   		OWF_Result[12].31:=0;
   	End_If;
   	If OWF_Input[5].[4] Then
   		OWF_Result[0]:=OWF_Result[0] + 1011754521+OWF_Add_c;
   		OWF_Add_c.0:=OWF_Result[0].31;
   		OWF_Result[0].31:=0;
   		OWF_Result[1]:=OWF_Result[1] + 1795510147+OWF_Add_c;
   		OWF_Add_c.1:=OWF_Result[1].31;
   		OWF_Result[1].31:=0;
   		OWF_Result[2]:=OWF_Result[2] + 543218634+OWF_Add_c;
   		OWF_Add_c.2:=OWF_Result[2].31;
   		OWF_Result[2].31:=0;
   		OWF_Result[3]:=OWF_Result[3] + 173475761+OWF_Add_c;
   		OWF_Add_c.3:=OWF_Result[3].31;
   		OWF_Result[3].31:=0;
   		OWF_Result[4]:=OWF_Result[4] + 535080772+OWF_Add_c;
   		OWF_Add_c.4:=OWF_Result[4].31;
   		OWF_Result[4].31:=0;
   		OWF_Result[5]:=OWF_Result[5] + 1289804735+OWF_Add_c;
   		OWF_Add_c.5:=OWF_Result[5].31;
   		OWF_Result[5].31:=0;
   		OWF_Result[6]:=OWF_Result[6] + 1812605489+OWF_Add_c;
   		OWF_Add_c.6:=OWF_Result[6].31;
   		OWF_Result[6].31:=0;
   		OWF_Result[7]:=OWF_Result[7] + 1203961891+OWF_Add_c;
   		OWF_Add_c.7:=OWF_Result[7].31;
   		OWF_Result[7].31:=0;
   		OWF_Result[8]:=OWF_Result[8] + 139150776+OWF_Add_c;
   		OWF_Add_c.8:=OWF_Result[8].31;
   		OWF_Result[8].31:=0;
   		OWF_Result[9]:=OWF_Result[9] + 1840895318+OWF_Add_c;
   		OWF_Add_c.9:=OWF_Result[9].31;
   		OWF_Result[9].31:=0;
   		OWF_Result[10]:=OWF_Result[10] + 576139644+OWF_Add_c;
   		OWF_Add_c.10:=OWF_Result[10].31;
   		OWF_Result[10].31:=0;
   		OWF_Result[11]:=OWF_Result[11] + 949700339+OWF_Add_c;
   		OWF_Add_c.11:=OWF_Result[11].31;
   		OWF_Result[11].31:=0;
   		OWF_Result[12]:=OWF_Result[12] + 707553602+OWF_Add_c;
   		OWF_Add_c.12:=OWF_Result[12].31;
   		OWF_Result[12].31:=0;
   	End_If;
   	If OWF_Input[5].[5] Then
   		OWF_Result[0]:=OWF_Result[0] + 341006670+OWF_Add_c;
   		OWF_Add_c.0:=OWF_Result[0].31;
   		OWF_Result[0].31:=0;
   		OWF_Result[1]:=OWF_Result[1] + 1545302097+OWF_Add_c;
   		OWF_Add_c.1:=OWF_Result[1].31;
   		OWF_Result[1].31:=0;
   		OWF_Result[2]:=OWF_Result[2] + 1059282447+OWF_Add_c;
   		OWF_Add_c.2:=OWF_Result[2].31;
   		OWF_Result[2].31:=0;
   		OWF_Result[3]:=OWF_Result[3] + 1918242377+OWF_Add_c;
   		OWF_Add_c.3:=OWF_Result[3].31;
   		OWF_Result[3].31:=0;
   		OWF_Result[4]:=OWF_Result[4] + 702854685+OWF_Add_c;
   		OWF_Add_c.4:=OWF_Result[4].31;
   		OWF_Result[4].31:=0;
   		OWF_Result[5]:=OWF_Result[5] + 1290612547+OWF_Add_c;
   		OWF_Add_c.5:=OWF_Result[5].31;
   		OWF_Result[5].31:=0;
   		OWF_Result[6]:=OWF_Result[6] + 1937985650+OWF_Add_c;
   		OWF_Add_c.6:=OWF_Result[6].31;
   		OWF_Result[6].31:=0;
   		OWF_Result[7]:=OWF_Result[7] + 1535904701+OWF_Add_c;
   		OWF_Add_c.7:=OWF_Result[7].31;
   		OWF_Result[7].31:=0;
   		OWF_Result[8]:=OWF_Result[8] + 57458357+OWF_Add_c;
   		OWF_Add_c.8:=OWF_Result[8].31;
   		OWF_Result[8].31:=0;
   		OWF_Result[9]:=OWF_Result[9] + 1270027244+OWF_Add_c;
   		OWF_Add_c.9:=OWF_Result[9].31;
   		OWF_Result[9].31:=0;
   		OWF_Result[10]:=OWF_Result[10] + 69146856+OWF_Add_c;
   		OWF_Add_c.10:=OWF_Result[10].31;
   		OWF_Result[10].31:=0;
   		OWF_Result[11]:=OWF_Result[11] + 1589075229+OWF_Add_c;
   		OWF_Add_c.11:=OWF_Result[11].31;
   		OWF_Result[11].31:=0;
   		OWF_Result[12]:=OWF_Result[12] + 458672961+OWF_Add_c;
   		OWF_Add_c.12:=OWF_Result[12].31;
   		OWF_Result[12].31:=0;
   	End_If;
   	If OWF_Input[5].[6] Then
   		OWF_Result[0]:=OWF_Result[0] + 1896310267+OWF_Add_c;
   		OWF_Add_c.0:=OWF_Result[0].31;
   		OWF_Result[0].31:=0;
   		OWF_Result[1]:=OWF_Result[1] + 1529180561+OWF_Add_c;
   		OWF_Add_c.1:=OWF_Result[1].31;
   		OWF_Result[1].31:=0;
   		OWF_Result[2]:=OWF_Result[2] + 2032481565+OWF_Add_c;
   		OWF_Add_c.2:=OWF_Result[2].31;
   		OWF_Result[2].31:=0;
   		OWF_Result[3]:=OWF_Result[3] + 537640111+OWF_Add_c;
   		OWF_Add_c.3:=OWF_Result[3].31;
   		OWF_Result[3].31:=0;
   		OWF_Result[4]:=OWF_Result[4] + 1272872794+OWF_Add_c;
   		OWF_Add_c.4:=OWF_Result[4].31;
   		OWF_Result[4].31:=0;
   		OWF_Result[5]:=OWF_Result[5] + 1539824454+OWF_Add_c;
   		OWF_Add_c.5:=OWF_Result[5].31;
   		OWF_Result[5].31:=0;
   		OWF_Result[6]:=OWF_Result[6] + 1430612137+OWF_Add_c;
   		OWF_Add_c.6:=OWF_Result[6].31;
   		OWF_Result[6].31:=0;
   		OWF_Result[7]:=OWF_Result[7] + 157560679+OWF_Add_c;
   		OWF_Add_c.7:=OWF_Result[7].31;
   		OWF_Result[7].31:=0;
   		OWF_Result[8]:=OWF_Result[8] + 259827156+OWF_Add_c;
   		OWF_Add_c.8:=OWF_Result[8].31;
   		OWF_Result[8].31:=0;
   		OWF_Result[9]:=OWF_Result[9] + 749936791+OWF_Add_c;
   		OWF_Add_c.9:=OWF_Result[9].31;
   		OWF_Result[9].31:=0;
   		OWF_Result[10]:=OWF_Result[10] + 1780248371+OWF_Add_c;
   		OWF_Add_c.10:=OWF_Result[10].31;
   		OWF_Result[10].31:=0;
   		OWF_Result[11]:=OWF_Result[11] + 1418315384+OWF_Add_c;
   		OWF_Add_c.11:=OWF_Result[11].31;
   		OWF_Result[11].31:=0;
   		OWF_Result[12]:=OWF_Result[12] + 406159660+OWF_Add_c;
   		OWF_Add_c.12:=OWF_Result[12].31;
   		OWF_Result[12].31:=0;
   	End_If;
   	If OWF_Input[5].[7] Then
   		OWF_Result[0]:=OWF_Result[0] + 2117716500+OWF_Add_c;
   		OWF_Add_c.0:=OWF_Result[0].31;
   		OWF_Result[0].31:=0;
   		OWF_Result[1]:=OWF_Result[1] + 1481111712+OWF_Add_c;
   		OWF_Add_c.1:=OWF_Result[1].31;
   		OWF_Result[1].31:=0;
   		OWF_Result[2]:=OWF_Result[2] + 1208238622+OWF_Add_c;
   		OWF_Add_c.2:=OWF_Result[2].31;
   		OWF_Result[2].31:=0;
   		OWF_Result[3]:=OWF_Result[3] + 1587378712+OWF_Add_c;
   		OWF_Add_c.3:=OWF_Result[3].31;
   		OWF_Result[3].31:=0;
   		OWF_Result[4]:=OWF_Result[4] + 1486187831+OWF_Add_c;
   		OWF_Add_c.4:=OWF_Result[4].31;
   		OWF_Result[4].31:=0;
   		OWF_Result[5]:=OWF_Result[5] + 1463632282+OWF_Add_c;
   		OWF_Add_c.5:=OWF_Result[5].31;
   		OWF_Result[5].31:=0;
   		OWF_Result[6]:=OWF_Result[6] + 594379430+OWF_Add_c;
   		OWF_Add_c.6:=OWF_Result[6].31;
   		OWF_Result[6].31:=0;
   		OWF_Result[7]:=OWF_Result[7] + 61907271+OWF_Add_c;
   		OWF_Add_c.7:=OWF_Result[7].31;
   		OWF_Result[7].31:=0;
   		OWF_Result[8]:=OWF_Result[8] + 1446292796+OWF_Add_c;
   		OWF_Add_c.8:=OWF_Result[8].31;
   		OWF_Result[8].31:=0;
   		OWF_Result[9]:=OWF_Result[9] + 1953507778+OWF_Add_c;
   		OWF_Add_c.9:=OWF_Result[9].31;
   		OWF_Result[9].31:=0;
   		OWF_Result[10]:=OWF_Result[10] + 1721398400+OWF_Add_c;
   		OWF_Add_c.10:=OWF_Result[10].31;
   		OWF_Result[10].31:=0;
   		OWF_Result[11]:=OWF_Result[11] + 704130819+OWF_Add_c;
   		OWF_Add_c.11:=OWF_Result[11].31;
   		OWF_Result[11].31:=0;
   		OWF_Result[12]:=OWF_Result[12] + 156099517+OWF_Add_c;
   		OWF_Add_c.12:=OWF_Result[12].31;
   		OWF_Result[12].31:=0;
   	End_If;
   	If OWF_Input[5].[8] Then
   		OWF_Result[0]:=OWF_Result[0] + 1443938657+OWF_Add_c;
   		OWF_Add_c.0:=OWF_Result[0].31;
   		OWF_Result[0].31:=0;
   		OWF_Result[1]:=OWF_Result[1] + 387077029+OWF_Add_c;
   		OWF_Add_c.1:=OWF_Result[1].31;
   		OWF_Result[1].31:=0;
   		OWF_Result[2]:=OWF_Result[2] + 331220417+OWF_Add_c;
   		OWF_Add_c.2:=OWF_Result[2].31;
   		OWF_Result[2].31:=0;
   		OWF_Result[3]:=OWF_Result[3] + 1153901105+OWF_Add_c;
   		OWF_Add_c.3:=OWF_Result[3].31;
   		OWF_Result[3].31:=0;
   		OWF_Result[4]:=OWF_Result[4] + 758718018+OWF_Add_c;
   		OWF_Add_c.4:=OWF_Result[4].31;
   		OWF_Result[4].31:=0;
   		OWF_Result[5]:=OWF_Result[5] + 1180469231+OWF_Add_c;
   		OWF_Add_c.5:=OWF_Result[5].31;
   		OWF_Result[5].31:=0;
   		OWF_Result[6]:=OWF_Result[6] + 451076221+OWF_Add_c;
   		OWF_Add_c.6:=OWF_Result[6].31;
   		OWF_Result[6].31:=0;
   		OWF_Result[7]:=OWF_Result[7] + 1957369555+OWF_Add_c;
   		OWF_Add_c.7:=OWF_Result[7].31;
   		OWF_Result[7].31:=0;
   		OWF_Result[8]:=OWF_Result[8] + 157679071+OWF_Add_c;
   		OWF_Add_c.8:=OWF_Result[8].31;
   		OWF_Result[8].31:=0;
   		OWF_Result[9]:=OWF_Result[9] + 999919265+OWF_Add_c;
   		OWF_Add_c.9:=OWF_Result[9].31;
   		OWF_Result[9].31:=0;
   		OWF_Result[10]:=OWF_Result[10] + 325782623+OWF_Add_c;
   		OWF_Add_c.10:=OWF_Result[10].31;
   		OWF_Result[10].31:=0;
   		OWF_Result[11]:=OWF_Result[11] + 1839549707+OWF_Add_c;
   		OWF_Add_c.11:=OWF_Result[11].31;
   		OWF_Result[11].31:=0;
   		OWF_Result[12]:=OWF_Result[12] + 210567637+OWF_Add_c;
   		OWF_Add_c.12:=OWF_Result[12].31;
   		OWF_Result[12].31:=0;
   	End_If;
   	If OWF_Input[5].[9] Then
   		OWF_Result[0]:=OWF_Result[0] + 1164800234+OWF_Add_c;
   		OWF_Add_c.0:=OWF_Result[0].31;
   		OWF_Result[0].31:=0;
   		OWF_Result[1]:=OWF_Result[1] + 373070247+OWF_Add_c;
   		OWF_Add_c.1:=OWF_Result[1].31;
   		OWF_Result[1].31:=0;
   		OWF_Result[2]:=OWF_Result[2] + 102655075+OWF_Add_c;
   		OWF_Add_c.2:=OWF_Result[2].31;
   		OWF_Result[2].31:=0;
   		OWF_Result[3]:=OWF_Result[3] + 1112504203+OWF_Add_c;
   		OWF_Add_c.3:=OWF_Result[3].31;
   		OWF_Result[3].31:=0;
   		OWF_Result[4]:=OWF_Result[4] + 728629506+OWF_Add_c;
   		OWF_Add_c.4:=OWF_Result[4].31;
   		OWF_Result[4].31:=0;
   		OWF_Result[5]:=OWF_Result[5] + 112310491+OWF_Add_c;
   		OWF_Add_c.5:=OWF_Result[5].31;
   		OWF_Result[5].31:=0;
   		OWF_Result[6]:=OWF_Result[6] + 1422404199+OWF_Add_c;
   		OWF_Add_c.6:=OWF_Result[6].31;
   		OWF_Result[6].31:=0;
   		OWF_Result[7]:=OWF_Result[7] + 1701166039+OWF_Add_c;
   		OWF_Add_c.7:=OWF_Result[7].31;
   		OWF_Result[7].31:=0;
   		OWF_Result[8]:=OWF_Result[8] + 2102782443+OWF_Add_c;
   		OWF_Add_c.8:=OWF_Result[8].31;
   		OWF_Result[8].31:=0;
   		OWF_Result[9]:=OWF_Result[9] + 1540134296+OWF_Add_c;
   		OWF_Add_c.9:=OWF_Result[9].31;
   		OWF_Result[9].31:=0;
   		OWF_Result[10]:=OWF_Result[10] + 2068205909+OWF_Add_c;
   		OWF_Add_c.10:=OWF_Result[10].31;
   		OWF_Result[10].31:=0;
   		OWF_Result[11]:=OWF_Result[11] + 1462437349+OWF_Add_c;
   		OWF_Add_c.11:=OWF_Result[11].31;
   		OWF_Result[11].31:=0;
   		OWF_Result[12]:=OWF_Result[12] + 1542204103+OWF_Add_c;
   		OWF_Add_c.12:=OWF_Result[12].31;
   		OWF_Result[12].31:=0;
   	End_If;
   	If OWF_Input[5].[10] Then
   		OWF_Result[0]:=OWF_Result[0] + 1094309781+OWF_Add_c;
   		OWF_Add_c.0:=OWF_Result[0].31;
   		OWF_Result[0].31:=0;
   		OWF_Result[1]:=OWF_Result[1] + 1799253283+OWF_Add_c;
   		OWF_Add_c.1:=OWF_Result[1].31;
   		OWF_Result[1].31:=0;
   		OWF_Result[2]:=OWF_Result[2] + 907784774+OWF_Add_c;
   		OWF_Add_c.2:=OWF_Result[2].31;
   		OWF_Result[2].31:=0;
   		OWF_Result[3]:=OWF_Result[3] + 1760595174+OWF_Add_c;
   		OWF_Add_c.3:=OWF_Result[3].31;
   		OWF_Result[3].31:=0;
   		OWF_Result[4]:=OWF_Result[4] + 1516380446+OWF_Add_c;
   		OWF_Add_c.4:=OWF_Result[4].31;
   		OWF_Result[4].31:=0;
   		OWF_Result[5]:=OWF_Result[5] + 525293244+OWF_Add_c;
   		OWF_Add_c.5:=OWF_Result[5].31;
   		OWF_Result[5].31:=0;
   		OWF_Result[6]:=OWF_Result[6] + 1469823607+OWF_Add_c;
   		OWF_Add_c.6:=OWF_Result[6].31;
   		OWF_Result[6].31:=0;
   		OWF_Result[7]:=OWF_Result[7] + 990094771+OWF_Add_c;
   		OWF_Add_c.7:=OWF_Result[7].31;
   		OWF_Result[7].31:=0;
   		OWF_Result[8]:=OWF_Result[8] + 206451193+OWF_Add_c;
   		OWF_Add_c.8:=OWF_Result[8].31;
   		OWF_Result[8].31:=0;
   		OWF_Result[9]:=OWF_Result[9] + 2094599626+OWF_Add_c;
   		OWF_Add_c.9:=OWF_Result[9].31;
   		OWF_Result[9].31:=0;
   		OWF_Result[10]:=OWF_Result[10] + 1804619518+OWF_Add_c;
   		OWF_Add_c.10:=OWF_Result[10].31;
   		OWF_Result[10].31:=0;
   		OWF_Result[11]:=OWF_Result[11] + 531327458+OWF_Add_c;
   		OWF_Add_c.11:=OWF_Result[11].31;
   		OWF_Result[11].31:=0;
   		OWF_Result[12]:=OWF_Result[12] + 914900243+OWF_Add_c;
   		OWF_Add_c.12:=OWF_Result[12].31;
   		OWF_Result[12].31:=0;
   	End_If;
   	If OWF_Input[5].[11] Then
   		OWF_Result[0]:=OWF_Result[0] + 1387671324+OWF_Add_c;
   		OWF_Add_c.0:=OWF_Result[0].31;
   		OWF_Result[0].31:=0;
   		OWF_Result[1]:=OWF_Result[1] + 770124107+OWF_Add_c;
   		OWF_Add_c.1:=OWF_Result[1].31;
   		OWF_Result[1].31:=0;
   		OWF_Result[2]:=OWF_Result[2] + 2104522684+OWF_Add_c;
   		OWF_Add_c.2:=OWF_Result[2].31;
   		OWF_Result[2].31:=0;
   		OWF_Result[3]:=OWF_Result[3] + 702616803+OWF_Add_c;
   		OWF_Add_c.3:=OWF_Result[3].31;
   		OWF_Result[3].31:=0;
   		OWF_Result[4]:=OWF_Result[4] + 453094356+OWF_Add_c;
   		OWF_Add_c.4:=OWF_Result[4].31;
   		OWF_Result[4].31:=0;
   		OWF_Result[5]:=OWF_Result[5] + 2109390133+OWF_Add_c;
   		OWF_Add_c.5:=OWF_Result[5].31;
   		OWF_Result[5].31:=0;
   		OWF_Result[6]:=OWF_Result[6] + 156781386+OWF_Add_c;
   		OWF_Add_c.6:=OWF_Result[6].31;
   		OWF_Result[6].31:=0;
   		OWF_Result[7]:=OWF_Result[7] + 1882451383+OWF_Add_c;
   		OWF_Add_c.7:=OWF_Result[7].31;
   		OWF_Result[7].31:=0;
   		OWF_Result[8]:=OWF_Result[8] + 1276007251+OWF_Add_c;
   		OWF_Add_c.8:=OWF_Result[8].31;
   		OWF_Result[8].31:=0;
   		OWF_Result[9]:=OWF_Result[9] + 1340635153+OWF_Add_c;
   		OWF_Add_c.9:=OWF_Result[9].31;
   		OWF_Result[9].31:=0;
   		OWF_Result[10]:=OWF_Result[10] + 225675392+OWF_Add_c;
   		OWF_Add_c.10:=OWF_Result[10].31;
   		OWF_Result[10].31:=0;
   		OWF_Result[11]:=OWF_Result[11] + 403241353+OWF_Add_c;
   		OWF_Add_c.11:=OWF_Result[11].31;
   		OWF_Result[11].31:=0;
   		OWF_Result[12]:=OWF_Result[12] + 1949018013+OWF_Add_c;
   		OWF_Add_c.12:=OWF_Result[12].31;
   		OWF_Result[12].31:=0;
   	End_If;
   	If OWF_Input[5].[12] Then
   		OWF_Result[0]:=OWF_Result[0] + 1384871639+OWF_Add_c;
   		OWF_Add_c.0:=OWF_Result[0].31;
   		OWF_Result[0].31:=0;
   		OWF_Result[1]:=OWF_Result[1] + 1594702713+OWF_Add_c;
   		OWF_Add_c.1:=OWF_Result[1].31;
   		OWF_Result[1].31:=0;
   		OWF_Result[2]:=OWF_Result[2] + 756803648+OWF_Add_c;
   		OWF_Add_c.2:=OWF_Result[2].31;
   		OWF_Result[2].31:=0;
   		OWF_Result[3]:=OWF_Result[3] + 26768879+OWF_Add_c;
   		OWF_Add_c.3:=OWF_Result[3].31;
   		OWF_Result[3].31:=0;
   		OWF_Result[4]:=OWF_Result[4] + 1679784822+OWF_Add_c;
   		OWF_Add_c.4:=OWF_Result[4].31;
   		OWF_Result[4].31:=0;
   		OWF_Result[5]:=OWF_Result[5] + 970059452+OWF_Add_c;
   		OWF_Add_c.5:=OWF_Result[5].31;
   		OWF_Result[5].31:=0;
   		OWF_Result[6]:=OWF_Result[6] + 1810393488+OWF_Add_c;
   		OWF_Add_c.6:=OWF_Result[6].31;
   		OWF_Result[6].31:=0;
   		OWF_Result[7]:=OWF_Result[7] + 488169811+OWF_Add_c;
   		OWF_Add_c.7:=OWF_Result[7].31;
   		OWF_Result[7].31:=0;
   		OWF_Result[8]:=OWF_Result[8] + 1304722861+OWF_Add_c;
   		OWF_Add_c.8:=OWF_Result[8].31;
   		OWF_Result[8].31:=0;
   		OWF_Result[9]:=OWF_Result[9] + 1892980786+OWF_Add_c;
   		OWF_Add_c.9:=OWF_Result[9].31;
   		OWF_Result[9].31:=0;
   		OWF_Result[10]:=OWF_Result[10] + 1092125948+OWF_Add_c;
   		OWF_Add_c.10:=OWF_Result[10].31;
   		OWF_Result[10].31:=0;
   		OWF_Result[11]:=OWF_Result[11] + 1982722541+OWF_Add_c;
   		OWF_Add_c.11:=OWF_Result[11].31;
   		OWF_Result[11].31:=0;
   		OWF_Result[12]:=OWF_Result[12] + 326633928+OWF_Add_c;
   		OWF_Add_c.12:=OWF_Result[12].31;
   		OWF_Result[12].31:=0;
   	End_If;
   	If OWF_Input[5].[13] Then
   		OWF_Result[0]:=OWF_Result[0] + 1000988417+OWF_Add_c;
   		OWF_Add_c.0:=OWF_Result[0].31;
   		OWF_Result[0].31:=0;
   		OWF_Result[1]:=OWF_Result[1] + 994193103+OWF_Add_c;
   		OWF_Add_c.1:=OWF_Result[1].31;
   		OWF_Result[1].31:=0;
   		OWF_Result[2]:=OWF_Result[2] + 1537710547+OWF_Add_c;
   		OWF_Add_c.2:=OWF_Result[2].31;
   		OWF_Result[2].31:=0;
   		OWF_Result[3]:=OWF_Result[3] + 15619081+OWF_Add_c;
   		OWF_Add_c.3:=OWF_Result[3].31;
   		OWF_Result[3].31:=0;
   		OWF_Result[4]:=OWF_Result[4] + 2143143663+OWF_Add_c;
   		OWF_Add_c.4:=OWF_Result[4].31;
   		OWF_Result[4].31:=0;
   		OWF_Result[5]:=OWF_Result[5] + 393950588+OWF_Add_c;
   		OWF_Add_c.5:=OWF_Result[5].31;
   		OWF_Result[5].31:=0;
   		OWF_Result[6]:=OWF_Result[6] + 1961783643+OWF_Add_c;
   		OWF_Add_c.6:=OWF_Result[6].31;
   		OWF_Result[6].31:=0;
   		OWF_Result[7]:=OWF_Result[7] + 2056947807+OWF_Add_c;
   		OWF_Add_c.7:=OWF_Result[7].31;
   		OWF_Result[7].31:=0;
   		OWF_Result[8]:=OWF_Result[8] + 939957448+OWF_Add_c;
   		OWF_Add_c.8:=OWF_Result[8].31;
   		OWF_Result[8].31:=0;
   		OWF_Result[9]:=OWF_Result[9] + 1853399300+OWF_Add_c;
   		OWF_Add_c.9:=OWF_Result[9].31;
   		OWF_Result[9].31:=0;
   		OWF_Result[10]:=OWF_Result[10] + 1339264557+OWF_Add_c;
   		OWF_Add_c.10:=OWF_Result[10].31;
   		OWF_Result[10].31:=0;
   		OWF_Result[11]:=OWF_Result[11] + 200481107+OWF_Add_c;
   		OWF_Add_c.11:=OWF_Result[11].31;
   		OWF_Result[11].31:=0;
   		OWF_Result[12]:=OWF_Result[12] + 1047995528+OWF_Add_c;
   		OWF_Add_c.12:=OWF_Result[12].31;
   		OWF_Result[12].31:=0;
   	End_If;
   	If OWF_Input[5].[14] Then
   		OWF_Result[0]:=OWF_Result[0] + 1208463242+OWF_Add_c;
   		OWF_Add_c.0:=OWF_Result[0].31;
   		OWF_Result[0].31:=0;
   		OWF_Result[1]:=OWF_Result[1] + 1623027587+OWF_Add_c;
   		OWF_Add_c.1:=OWF_Result[1].31;
   		OWF_Result[1].31:=0;
   		OWF_Result[2]:=OWF_Result[2] + 605083722+OWF_Add_c;
   		OWF_Add_c.2:=OWF_Result[2].31;
   		OWF_Result[2].31:=0;
   		OWF_Result[3]:=OWF_Result[3] + 1196976689+OWF_Add_c;
   		OWF_Add_c.3:=OWF_Result[3].31;
   		OWF_Result[3].31:=0;
   		OWF_Result[4]:=OWF_Result[4] + 2034493170+OWF_Add_c;
   		OWF_Add_c.4:=OWF_Result[4].31;
   		OWF_Result[4].31:=0;
   		OWF_Result[5]:=OWF_Result[5] + 718055369+OWF_Add_c;
   		OWF_Add_c.5:=OWF_Result[5].31;
   		OWF_Result[5].31:=0;
   		OWF_Result[6]:=OWF_Result[6] + 910332765+OWF_Add_c;
   		OWF_Add_c.6:=OWF_Result[6].31;
   		OWF_Result[6].31:=0;
   		OWF_Result[7]:=OWF_Result[7] + 1449925077+OWF_Add_c;
   		OWF_Add_c.7:=OWF_Result[7].31;
   		OWF_Result[7].31:=0;
   		OWF_Result[8]:=OWF_Result[8] + 839039994+OWF_Add_c;
   		OWF_Add_c.8:=OWF_Result[8].31;
   		OWF_Result[8].31:=0;
   		OWF_Result[9]:=OWF_Result[9] + 1168597276+OWF_Add_c;
   		OWF_Add_c.9:=OWF_Result[9].31;
   		OWF_Result[9].31:=0;
   		OWF_Result[10]:=OWF_Result[10] + 42917457+OWF_Add_c;
   		OWF_Add_c.10:=OWF_Result[10].31;
   		OWF_Result[10].31:=0;
   		OWF_Result[11]:=OWF_Result[11] + 1907752552+OWF_Add_c;
   		OWF_Add_c.11:=OWF_Result[11].31;
   		OWF_Result[11].31:=0;
   		OWF_Result[12]:=OWF_Result[12] + 1741695515+OWF_Add_c;
   		OWF_Add_c.12:=OWF_Result[12].31;
   		OWF_Result[12].31:=0;
   	End_If;
   	If OWF_Input[5].[15] Then
   		OWF_Result[0]:=OWF_Result[0] + 963845262+OWF_Add_c;
   		OWF_Add_c.0:=OWF_Result[0].31;
   		OWF_Result[0].31:=0;
   		OWF_Result[1]:=OWF_Result[1] + 1178480242+OWF_Add_c;
   		OWF_Add_c.1:=OWF_Result[1].31;
   		OWF_Result[1].31:=0;
   		OWF_Result[2]:=OWF_Result[2] + 555963648+OWF_Add_c;
   		OWF_Add_c.2:=OWF_Result[2].31;
   		OWF_Result[2].31:=0;
   		OWF_Result[3]:=OWF_Result[3] + 2035289100+OWF_Add_c;
   		OWF_Add_c.3:=OWF_Result[3].31;
   		OWF_Result[3].31:=0;
   		OWF_Result[4]:=OWF_Result[4] + 1602592723+OWF_Add_c;
   		OWF_Add_c.4:=OWF_Result[4].31;
   		OWF_Result[4].31:=0;
   		OWF_Result[5]:=OWF_Result[5] + 1321176695+OWF_Add_c;
   		OWF_Add_c.5:=OWF_Result[5].31;
   		OWF_Result[5].31:=0;
   		OWF_Result[6]:=OWF_Result[6] + 1370169932+OWF_Add_c;
   		OWF_Add_c.6:=OWF_Result[6].31;
   		OWF_Result[6].31:=0;
   		OWF_Result[7]:=OWF_Result[7] + 1543393295+OWF_Add_c;
   		OWF_Add_c.7:=OWF_Result[7].31;
   		OWF_Result[7].31:=0;
   		OWF_Result[8]:=OWF_Result[8] + 83738279+OWF_Add_c;
   		OWF_Add_c.8:=OWF_Result[8].31;
   		OWF_Result[8].31:=0;
   		OWF_Result[9]:=OWF_Result[9] + 725427957+OWF_Add_c;
   		OWF_Add_c.9:=OWF_Result[9].31;
   		OWF_Result[9].31:=0;
   		OWF_Result[10]:=OWF_Result[10] + 581206308+OWF_Add_c;
   		OWF_Add_c.10:=OWF_Result[10].31;
   		OWF_Result[10].31:=0;
   		OWF_Result[11]:=OWF_Result[11] + 491262647+OWF_Add_c;
   		OWF_Add_c.11:=OWF_Result[11].31;
   		OWF_Result[11].31:=0;
   		OWF_Result[12]:=OWF_Result[12] + 2147137437+OWF_Add_c;
   		OWF_Add_c.12:=OWF_Result[12].31;
   		OWF_Result[12].31:=0;
   	End_If;
   	If OWF_Input[5].[16] Then
   		OWF_Result[0]:=OWF_Result[0] + 2074453075+OWF_Add_c;
   		OWF_Add_c.0:=OWF_Result[0].31;
   		OWF_Result[0].31:=0;
   		OWF_Result[1]:=OWF_Result[1] + 108344464+OWF_Add_c;
   		OWF_Add_c.1:=OWF_Result[1].31;
   		OWF_Result[1].31:=0;
   		OWF_Result[2]:=OWF_Result[2] + 452532141+OWF_Add_c;
   		OWF_Add_c.2:=OWF_Result[2].31;
   		OWF_Result[2].31:=0;
   		OWF_Result[3]:=OWF_Result[3] + 1547961836+OWF_Add_c;
   		OWF_Add_c.3:=OWF_Result[3].31;
   		OWF_Result[3].31:=0;
   		OWF_Result[4]:=OWF_Result[4] + 1372224157+OWF_Add_c;
   		OWF_Add_c.4:=OWF_Result[4].31;
   		OWF_Result[4].31:=0;
   		OWF_Result[5]:=OWF_Result[5] + 1842815326+OWF_Add_c;
   		OWF_Add_c.5:=OWF_Result[5].31;
   		OWF_Result[5].31:=0;
   		OWF_Result[6]:=OWF_Result[6] + 614084210+OWF_Add_c;
   		OWF_Add_c.6:=OWF_Result[6].31;
   		OWF_Result[6].31:=0;
   		OWF_Result[7]:=OWF_Result[7] + 2105622125+OWF_Add_c;
   		OWF_Add_c.7:=OWF_Result[7].31;
   		OWF_Result[7].31:=0;
   		OWF_Result[8]:=OWF_Result[8] + 1347171274+OWF_Add_c;
   		OWF_Add_c.8:=OWF_Result[8].31;
   		OWF_Result[8].31:=0;
   		OWF_Result[9]:=OWF_Result[9] + 1124490238+OWF_Add_c;
   		OWF_Add_c.9:=OWF_Result[9].31;
   		OWF_Result[9].31:=0;
   		OWF_Result[10]:=OWF_Result[10] + 2064336718+OWF_Add_c;
   		OWF_Add_c.10:=OWF_Result[10].31;
   		OWF_Result[10].31:=0;
   		OWF_Result[11]:=OWF_Result[11] + 1049919562+OWF_Add_c;
   		OWF_Add_c.11:=OWF_Result[11].31;
   		OWF_Result[11].31:=0;
   		OWF_Result[12]:=OWF_Result[12] + 13830202+OWF_Add_c;
   		OWF_Add_c.12:=OWF_Result[12].31;
   		OWF_Result[12].31:=0;
   	End_If;
   	If OWF_Input[5].[17] Then
   		OWF_Result[0]:=OWF_Result[0] + 409887176+OWF_Add_c;
   		OWF_Add_c.0:=OWF_Result[0].31;
   		OWF_Result[0].31:=0;
   		OWF_Result[1]:=OWF_Result[1] + 317844364+OWF_Add_c;
   		OWF_Add_c.1:=OWF_Result[1].31;
   		OWF_Result[1].31:=0;
   		OWF_Result[2]:=OWF_Result[2] + 232272628+OWF_Add_c;
   		OWF_Add_c.2:=OWF_Result[2].31;
   		OWF_Result[2].31:=0;
   		OWF_Result[3]:=OWF_Result[3] + 284187670+OWF_Add_c;
   		OWF_Add_c.3:=OWF_Result[3].31;
   		OWF_Result[3].31:=0;
   		OWF_Result[4]:=OWF_Result[4] + 1431286202+OWF_Add_c;
   		OWF_Add_c.4:=OWF_Result[4].31;
   		OWF_Result[4].31:=0;
   		OWF_Result[5]:=OWF_Result[5] + 1935493368+OWF_Add_c;
   		OWF_Add_c.5:=OWF_Result[5].31;
   		OWF_Result[5].31:=0;
   		OWF_Result[6]:=OWF_Result[6] + 1179830512+OWF_Add_c;
   		OWF_Add_c.6:=OWF_Result[6].31;
   		OWF_Result[6].31:=0;
   		OWF_Result[7]:=OWF_Result[7] + 553237340+OWF_Add_c;
   		OWF_Add_c.7:=OWF_Result[7].31;
   		OWF_Result[7].31:=0;
   		OWF_Result[8]:=OWF_Result[8] + 374481235+OWF_Add_c;
   		OWF_Add_c.8:=OWF_Result[8].31;
   		OWF_Result[8].31:=0;
   		OWF_Result[9]:=OWF_Result[9] + 699596432+OWF_Add_c;
   		OWF_Add_c.9:=OWF_Result[9].31;
   		OWF_Result[9].31:=0;
   		OWF_Result[10]:=OWF_Result[10] + 1347480733+OWF_Add_c;
   		OWF_Add_c.10:=OWF_Result[10].31;
   		OWF_Result[10].31:=0;
   		OWF_Result[11]:=OWF_Result[11] + 867993303+OWF_Add_c;
   		OWF_Add_c.11:=OWF_Result[11].31;
   		OWF_Result[11].31:=0;
   		OWF_Result[12]:=OWF_Result[12] + 1741665324+OWF_Add_c;
   		OWF_Add_c.12:=OWF_Result[12].31;
   		OWF_Result[12].31:=0;
   	End_If;
   	If OWF_Input[5].[18] Then
   		OWF_Result[0]:=OWF_Result[0] + 181112595+OWF_Add_c;
   		OWF_Add_c.0:=OWF_Result[0].31;
   		OWF_Result[0].31:=0;
   		OWF_Result[1]:=OWF_Result[1] + 1763223656+OWF_Add_c;
   		OWF_Add_c.1:=OWF_Result[1].31;
   		OWF_Result[1].31:=0;
   		OWF_Result[2]:=OWF_Result[2] + 228534745+OWF_Add_c;
   		OWF_Add_c.2:=OWF_Result[2].31;
   		OWF_Result[2].31:=0;
   		OWF_Result[3]:=OWF_Result[3] + 1241484761+OWF_Add_c;
   		OWF_Add_c.3:=OWF_Result[3].31;
   		OWF_Result[3].31:=0;
   		OWF_Result[4]:=OWF_Result[4] + 2081376218+OWF_Add_c;
   		OWF_Add_c.4:=OWF_Result[4].31;
   		OWF_Result[4].31:=0;
   		OWF_Result[5]:=OWF_Result[5] + 883325201+OWF_Add_c;
   		OWF_Add_c.5:=OWF_Result[5].31;
   		OWF_Result[5].31:=0;
   		OWF_Result[6]:=OWF_Result[6] + 1084382409+OWF_Add_c;
   		OWF_Add_c.6:=OWF_Result[6].31;
   		OWF_Result[6].31:=0;
   		OWF_Result[7]:=OWF_Result[7] + 810849280+OWF_Add_c;
   		OWF_Add_c.7:=OWF_Result[7].31;
   		OWF_Result[7].31:=0;
   		OWF_Result[8]:=OWF_Result[8] + 1583250563+OWF_Add_c;
   		OWF_Add_c.8:=OWF_Result[8].31;
   		OWF_Result[8].31:=0;
   		OWF_Result[9]:=OWF_Result[9] + 234577571+OWF_Add_c;
   		OWF_Add_c.9:=OWF_Result[9].31;
   		OWF_Result[9].31:=0;
   		OWF_Result[10]:=OWF_Result[10] + 1030400922+OWF_Add_c;
   		OWF_Add_c.10:=OWF_Result[10].31;
   		OWF_Result[10].31:=0;
   		OWF_Result[11]:=OWF_Result[11] + 746653471+OWF_Add_c;
   		OWF_Add_c.11:=OWF_Result[11].31;
   		OWF_Result[11].31:=0;
   		OWF_Result[12]:=OWF_Result[12] + 1862214324+OWF_Add_c;
   		OWF_Add_c.12:=OWF_Result[12].31;
   		OWF_Result[12].31:=0;
   	End_If;
   	If OWF_Input[5].[19] Then
   		OWF_Result[0]:=OWF_Result[0] + 905287854+OWF_Add_c;
   		OWF_Add_c.0:=OWF_Result[0].31;
   		OWF_Result[0].31:=0;
   		OWF_Result[1]:=OWF_Result[1] + 171069296+OWF_Add_c;
   		OWF_Add_c.1:=OWF_Result[1].31;
   		OWF_Result[1].31:=0;
   		OWF_Result[2]:=OWF_Result[2] + 922090179+OWF_Add_c;
   		OWF_Add_c.2:=OWF_Result[2].31;
   		OWF_Result[2].31:=0;
   		OWF_Result[3]:=OWF_Result[3] + 1913120820+OWF_Add_c;
   		OWF_Add_c.3:=OWF_Result[3].31;
   		OWF_Result[3].31:=0;
   		OWF_Result[4]:=OWF_Result[4] + 1248967781+OWF_Add_c;
   		OWF_Add_c.4:=OWF_Result[4].31;
   		OWF_Result[4].31:=0;
   		OWF_Result[5]:=OWF_Result[5] + 2027397171+OWF_Add_c;
   		OWF_Add_c.5:=OWF_Result[5].31;
   		OWF_Result[5].31:=0;
   		OWF_Result[6]:=OWF_Result[6] + 1771258503+OWF_Add_c;
   		OWF_Add_c.6:=OWF_Result[6].31;
   		OWF_Result[6].31:=0;
   		OWF_Result[7]:=OWF_Result[7] + 1286847095+OWF_Add_c;
   		OWF_Add_c.7:=OWF_Result[7].31;
   		OWF_Result[7].31:=0;
   		OWF_Result[8]:=OWF_Result[8] + 631683880+OWF_Add_c;
   		OWF_Add_c.8:=OWF_Result[8].31;
   		OWF_Result[8].31:=0;
   		OWF_Result[9]:=OWF_Result[9] + 1930526467+OWF_Add_c;
   		OWF_Add_c.9:=OWF_Result[9].31;
   		OWF_Result[9].31:=0;
   		OWF_Result[10]:=OWF_Result[10] + 844525456+OWF_Add_c;
   		OWF_Add_c.10:=OWF_Result[10].31;
   		OWF_Result[10].31:=0;
   		OWF_Result[11]:=OWF_Result[11] + 76605356+OWF_Add_c;
   		OWF_Add_c.11:=OWF_Result[11].31;
   		OWF_Result[11].31:=0;
   		OWF_Result[12]:=OWF_Result[12] + 1240692862+OWF_Add_c;
   		OWF_Add_c.12:=OWF_Result[12].31;
   		OWF_Result[12].31:=0;
   	End_If;
   	If OWF_Input[5].[20] Then
   		OWF_Result[0]:=OWF_Result[0] + 947806239+OWF_Add_c;
   		OWF_Add_c.0:=OWF_Result[0].31;
   		OWF_Result[0].31:=0;
   		OWF_Result[1]:=OWF_Result[1] + 1809109131+OWF_Add_c;
   		OWF_Add_c.1:=OWF_Result[1].31;
   		OWF_Result[1].31:=0;
   		OWF_Result[2]:=OWF_Result[2] + 353300745+OWF_Add_c;
   		OWF_Add_c.2:=OWF_Result[2].31;
   		OWF_Result[2].31:=0;
   		OWF_Result[3]:=OWF_Result[3] + 1824622451+OWF_Add_c;
   		OWF_Add_c.3:=OWF_Result[3].31;
   		OWF_Result[3].31:=0;
   		OWF_Result[4]:=OWF_Result[4] + 1679263964+OWF_Add_c;
   		OWF_Add_c.4:=OWF_Result[4].31;
   		OWF_Result[4].31:=0;
   		OWF_Result[5]:=OWF_Result[5] + 406258292+OWF_Add_c;
   		OWF_Add_c.5:=OWF_Result[5].31;
   		OWF_Result[5].31:=0;
   		OWF_Result[6]:=OWF_Result[6] + 1136140073+OWF_Add_c;
   		OWF_Add_c.6:=OWF_Result[6].31;
   		OWF_Result[6].31:=0;
   		OWF_Result[7]:=OWF_Result[7] + 320216123+OWF_Add_c;
   		OWF_Add_c.7:=OWF_Result[7].31;
   		OWF_Result[7].31:=0;
   		OWF_Result[8]:=OWF_Result[8] + 1349498735+OWF_Add_c;
   		OWF_Add_c.8:=OWF_Result[8].31;
   		OWF_Result[8].31:=0;
   		OWF_Result[9]:=OWF_Result[9] + 1095559942+OWF_Add_c;
   		OWF_Add_c.9:=OWF_Result[9].31;
   		OWF_Result[9].31:=0;
   		OWF_Result[10]:=OWF_Result[10] + 1701678166+OWF_Add_c;
   		OWF_Add_c.10:=OWF_Result[10].31;
   		OWF_Result[10].31:=0;
   		OWF_Result[11]:=OWF_Result[11] + 1167402895+OWF_Add_c;
   		OWF_Add_c.11:=OWF_Result[11].31;
   		OWF_Result[11].31:=0;
   		OWF_Result[12]:=OWF_Result[12] + 396826993+OWF_Add_c;
   		OWF_Add_c.12:=OWF_Result[12].31;
   		OWF_Result[12].31:=0;
   	End_If;
   	If OWF_Input[5].[21] Then
   		OWF_Result[0]:=OWF_Result[0] + 1459274711+OWF_Add_c;
   		OWF_Add_c.0:=OWF_Result[0].31;
   		OWF_Result[0].31:=0;
   		OWF_Result[1]:=OWF_Result[1] + 1739394073+OWF_Add_c;
   		OWF_Add_c.1:=OWF_Result[1].31;
   		OWF_Result[1].31:=0;
   		OWF_Result[2]:=OWF_Result[2] + 311010767+OWF_Add_c;
   		OWF_Add_c.2:=OWF_Result[2].31;
   		OWF_Result[2].31:=0;
   		OWF_Result[3]:=OWF_Result[3] + 226622081+OWF_Add_c;
   		OWF_Add_c.3:=OWF_Result[3].31;
   		OWF_Result[3].31:=0;
   		OWF_Result[4]:=OWF_Result[4] + 1368798677+OWF_Add_c;
   		OWF_Add_c.4:=OWF_Result[4].31;
   		OWF_Result[4].31:=0;
   		OWF_Result[5]:=OWF_Result[5] + 325030175+OWF_Add_c;
   		OWF_Add_c.5:=OWF_Result[5].31;
   		OWF_Result[5].31:=0;
   		OWF_Result[6]:=OWF_Result[6] + 1557429054+OWF_Add_c;
   		OWF_Add_c.6:=OWF_Result[6].31;
   		OWF_Result[6].31:=0;
   		OWF_Result[7]:=OWF_Result[7] + 312683037+OWF_Add_c;
   		OWF_Add_c.7:=OWF_Result[7].31;
   		OWF_Result[7].31:=0;
   		OWF_Result[8]:=OWF_Result[8] + 1059027382+OWF_Add_c;
   		OWF_Add_c.8:=OWF_Result[8].31;
   		OWF_Result[8].31:=0;
   		OWF_Result[9]:=OWF_Result[9] + 539763246+OWF_Add_c;
   		OWF_Add_c.9:=OWF_Result[9].31;
   		OWF_Result[9].31:=0;
   		OWF_Result[10]:=OWF_Result[10] + 380927532+OWF_Add_c;
   		OWF_Add_c.10:=OWF_Result[10].31;
   		OWF_Result[10].31:=0;
   		OWF_Result[11]:=OWF_Result[11] + 2033647151+OWF_Add_c;
   		OWF_Add_c.11:=OWF_Result[11].31;
   		OWF_Result[11].31:=0;
   		OWF_Result[12]:=OWF_Result[12] + 1263432976+OWF_Add_c;
   		OWF_Add_c.12:=OWF_Result[12].31;
   		OWF_Result[12].31:=0;
   	End_If;
   	If OWF_Input[5].[22] Then
   		OWF_Result[0]:=OWF_Result[0] + 850490276+OWF_Add_c;
   		OWF_Add_c.0:=OWF_Result[0].31;
   		OWF_Result[0].31:=0;
   		OWF_Result[1]:=OWF_Result[1] + 1505434702+OWF_Add_c;
   		OWF_Add_c.1:=OWF_Result[1].31;
   		OWF_Result[1].31:=0;
   		OWF_Result[2]:=OWF_Result[2] + 1435880615+OWF_Add_c;
   		OWF_Add_c.2:=OWF_Result[2].31;
   		OWF_Result[2].31:=0;
   		OWF_Result[3]:=OWF_Result[3] + 757815124+OWF_Add_c;
   		OWF_Add_c.3:=OWF_Result[3].31;
   		OWF_Result[3].31:=0;
   		OWF_Result[4]:=OWF_Result[4] + 226106502+OWF_Add_c;
   		OWF_Add_c.4:=OWF_Result[4].31;
   		OWF_Result[4].31:=0;
   		OWF_Result[5]:=OWF_Result[5] + 382560411+OWF_Add_c;
   		OWF_Add_c.5:=OWF_Result[5].31;
   		OWF_Result[5].31:=0;
   		OWF_Result[6]:=OWF_Result[6] + 1080056679+OWF_Add_c;
   		OWF_Add_c.6:=OWF_Result[6].31;
   		OWF_Result[6].31:=0;
   		OWF_Result[7]:=OWF_Result[7] + 20127395+OWF_Add_c;
   		OWF_Add_c.7:=OWF_Result[7].31;
   		OWF_Result[7].31:=0;
   		OWF_Result[8]:=OWF_Result[8] + 1148820067+OWF_Add_c;
   		OWF_Add_c.8:=OWF_Result[8].31;
   		OWF_Result[8].31:=0;
   		OWF_Result[9]:=OWF_Result[9] + 924116637+OWF_Add_c;
   		OWF_Add_c.9:=OWF_Result[9].31;
   		OWF_Result[9].31:=0;
   		OWF_Result[10]:=OWF_Result[10] + 676425310+OWF_Add_c;
   		OWF_Add_c.10:=OWF_Result[10].31;
   		OWF_Result[10].31:=0;
   		OWF_Result[11]:=OWF_Result[11] + 488537624+OWF_Add_c;
   		OWF_Add_c.11:=OWF_Result[11].31;
   		OWF_Result[11].31:=0;
   		OWF_Result[12]:=OWF_Result[12] + 1095846979+OWF_Add_c;
   		OWF_Add_c.12:=OWF_Result[12].31;
   		OWF_Result[12].31:=0;
   	End_If;
   	If OWF_Input[5].[23] Then
   		OWF_Result[0]:=OWF_Result[0] + 2136207919+OWF_Add_c;
   		OWF_Add_c.0:=OWF_Result[0].31;
   		OWF_Result[0].31:=0;
   		OWF_Result[1]:=OWF_Result[1] + 1736056703+OWF_Add_c;
   		OWF_Add_c.1:=OWF_Result[1].31;
   		OWF_Result[1].31:=0;
   		OWF_Result[2]:=OWF_Result[2] + 541452115+OWF_Add_c;
   		OWF_Add_c.2:=OWF_Result[2].31;
   		OWF_Result[2].31:=0;
   		OWF_Result[3]:=OWF_Result[3] + 1819467400+OWF_Add_c;
   		OWF_Add_c.3:=OWF_Result[3].31;
   		OWF_Result[3].31:=0;
   		OWF_Result[4]:=OWF_Result[4] + 1089042793+OWF_Add_c;
   		OWF_Add_c.4:=OWF_Result[4].31;
   		OWF_Result[4].31:=0;
   		OWF_Result[5]:=OWF_Result[5] + 800641240+OWF_Add_c;
   		OWF_Add_c.5:=OWF_Result[5].31;
   		OWF_Result[5].31:=0;
   		OWF_Result[6]:=OWF_Result[6] + 1848283435+OWF_Add_c;
   		OWF_Add_c.6:=OWF_Result[6].31;
   		OWF_Result[6].31:=0;
   		OWF_Result[7]:=OWF_Result[7] + 768914757+OWF_Add_c;
   		OWF_Add_c.7:=OWF_Result[7].31;
   		OWF_Result[7].31:=0;
   		OWF_Result[8]:=OWF_Result[8] + 1703211083+OWF_Add_c;
   		OWF_Add_c.8:=OWF_Result[8].31;
   		OWF_Result[8].31:=0;
   		OWF_Result[9]:=OWF_Result[9] + 1652863001+OWF_Add_c;
   		OWF_Add_c.9:=OWF_Result[9].31;
   		OWF_Result[9].31:=0;
   		OWF_Result[10]:=OWF_Result[10] + 1426503011+OWF_Add_c;
   		OWF_Add_c.10:=OWF_Result[10].31;
   		OWF_Result[10].31:=0;
   		OWF_Result[11]:=OWF_Result[11] + 237171419+OWF_Add_c;
   		OWF_Add_c.11:=OWF_Result[11].31;
   		OWF_Result[11].31:=0;
   		OWF_Result[12]:=OWF_Result[12] + 647871692+OWF_Add_c;
   		OWF_Add_c.12:=OWF_Result[12].31;
   		OWF_Result[12].31:=0;
   	End_If;
   	If OWF_Input[5].[24] Then
   		OWF_Result[0]:=OWF_Result[0] + 1463455914+OWF_Add_c;
   		OWF_Add_c.0:=OWF_Result[0].31;
   		OWF_Result[0].31:=0;
   		OWF_Result[1]:=OWF_Result[1] + 1733152448+OWF_Add_c;
   		OWF_Add_c.1:=OWF_Result[1].31;
   		OWF_Result[1].31:=0;
   		OWF_Result[2]:=OWF_Result[2] + 513694058+OWF_Add_c;
   		OWF_Add_c.2:=OWF_Result[2].31;
   		OWF_Result[2].31:=0;
   		OWF_Result[3]:=OWF_Result[3] + 2049031827+OWF_Add_c;
   		OWF_Add_c.3:=OWF_Result[3].31;
   		OWF_Result[3].31:=0;
   		OWF_Result[4]:=OWF_Result[4] + 571902437+OWF_Add_c;
   		OWF_Add_c.4:=OWF_Result[4].31;
   		OWF_Result[4].31:=0;
   		OWF_Result[5]:=OWF_Result[5] + 213654157+OWF_Add_c;
   		OWF_Add_c.5:=OWF_Result[5].31;
   		OWF_Result[5].31:=0;
   		OWF_Result[6]:=OWF_Result[6] + 1187052200+OWF_Add_c;
